
screen "02 Wip Select" 480x800, template "Current Menu Selection"
   Button "Top" at 375,164 size 100x101; TextOff 'Text'; PictureOff "basic panel top"
      on Press: function_b14e0dd5("pbs", 0)
      Appearance <- "[0]"
      Visibility <- "[0]"
   Button "Page Up" at 375,270 size 100x101; TextOff 'Text'; PictureOff "basic panel page up"
      on Press: function_b14e0dd5("pbs", 1)
      Visibility <- "[1]"
      Appearance <- "[1]"
   Button "Line Up" at 375,376 size 100x101; TextOff 'Text'; PictureOff "basic panel line up"
      on Press: function_b14e0dd5("pbs", 2)
      Appearance <- "[2]"
      Visibility <- "[2]"
   Button "Line Down" at 375,482 size 100x101; TextOff 'Text'; PictureOff "basic panel line down"
      on Press: function_b14e0dd5("pbs", 3)
      Visibility <- "[3]"
      Appearance <- "[3]"
   Button "Page Down" at 375,588 size 100x101; TextOff 'Text'; PictureOff "basic panel page down"
      on Press: function_b14e0dd5("pbs", 4)
      Appearance <- "[4]"
      Visibility <- "[4]"
   Button "Bottom" at 375,694 size 100x101; TextOff 'Text'; PictureOff "basic panel bottom"
      on Press: function_b14e0dd5("pbs", 5)
      Visibility <- "[5]"
      Appearance <- "[5]"
   IOField "brdrShortR00" at 5,164 size 365x101; FormatPattern 1
      Visibility <- "[6]"
      Appearance <- "[6]"
   IOField "brdrShortR01" at 5,270 size 365x101; FormatPattern 1
      Visibility <- "[7]"
      Appearance <- "[7]"
   IOField "brdrShortR02" at 5,376 size 365x101; FormatPattern 1
      Visibility <- "[8]"
      Appearance <- "[8]"
   IOField "brdrShortR03" at 5,482 size 365x101; FormatPattern 1
      Visibility <- "[9]"
      Appearance <- "[9]"
   IOField "brdrShortR04" at 5,588 size 365x101; FormatPattern 1
      Visibility <- "[10]"
      Appearance <- "[10]"
   IOField "brdrShortR05" at 5,694 size 365x101; FormatPattern 1
      Visibility <- "[11]"
      Appearance <- "[11]"
   Button "pbShortSelectR00" at 5,164 size 365x101; TextOff 'Text'
      on Release: ActivateScreen("01 Part Select", 0)
      on Press: function_b14e0dd5("pbs", 6)
   Button "pbShortSelectR01" at 5,270 size 365x101; TextOff 'Text'
      on Release: ActivateScreen("01 Part Select", 0)
      on Press: function_b14e0dd5("pbs", 7)
   Button "pbShortSelectR02" at 5,376 size 365x101; TextOff 'Text'
      on Release: ActivateScreen("01 Part Select", 0)
      on Press: function_b14e0dd5("pbs", 8)
   Button "pbShortSelectR03" at 5,482 size 365x101; TextOff 'Text'
      on Release: ActivateScreen("01 Part Select", 0)
      on Press: function_b14e0dd5("pbs", 9)
   Button "pbShortSelectR04" at 5,588 size 365x101; TextOff 'Text'
      on Release: ActivateScreen("01 Part Select", 0)
      on Press: function_b14e0dd5("pbs", 10)
   Button "pbShortSelectR05" at 5,694 size 365x101; TextOff 'Text'
      on Release: ActivateScreen("01 Part Select", 0)
      on Press: function_b14e0dd5("pbs", 11)
   IOField "brdrLongR00" at 5,164 size 470x101; FormatPattern 1
      Visibility <- "[18]"
   IOField "brdrLongR01" at 5,270 size 470x101; FormatPattern 1
      Visibility <- "[19]"
   IOField "brdrLongR02" at 5,376 size 470x101; FormatPattern 1
      Visibility <- "[20]"
   IOField "brdrLongR03" at 5,482 size 470x101; FormatPattern 1
      Visibility <- "[21]"
   IOField "brdrLongR04" at 5,588 size 470x101; FormatPattern 1
      Visibility <- "[22]"
   IOField "brdrLongR05" at 5,694 size 470x101; FormatPattern 1
      Visibility <- "[23]"
   Button "pbLongtSelectR00" at 5,164 size 470x101; TextOff 'Text'
      on Release: ActivateScreen("01 Part Select", 0)
      on Press: function_b14e0dd5("pbs", 6)
      Visibility <- "[18]"
   Button "pbLongtSelectR01" at 5,270 size 470x101; TextOff 'Text'
      on Release: ActivateScreen("01 Part Select", 0)
      on Press: function_b14e0dd5("pbs", 7)
      Visibility <- "[19]"
   Button "pbLongtSelectR02" at 5,376 size 470x101; TextOff 'Text'
      on Release: ActivateScreen("01 Part Select", 0)
      on Press: function_b14e0dd5("pbs", 8)
      Visibility <- "[20]"
   Button "pbLongtSelectR03" at 5,482 size 470x101; TextOff 'Text'
      on Release: ActivateScreen("01 Part Select", 0)
      on Press: function_b14e0dd5("pbs", 9)
      Visibility <- "[21]"
   Button "pbLongtSelectR04" at 5,588 size 470x101; TextOff 'Text'
      on Release: ActivateScreen("01 Part Select", 0)
      on Press: function_b14e0dd5("pbs", 10)
      Visibility <- "[22]"
   Button "pbLongtSelectR05" at 5,694 size 470x101; TextOff 'Text'
      on Release: ActivateScreen("01 Part Select", 0)
      on Press: function_b14e0dd5("pbs", 11)
      Visibility <- "[23]"
   IOField "iofLongtMenuSelectR00" at 42,166 size 430x97; FormatPattern ????????????????????????????????????????????????????????????
      Visibility <- "[18]"
      Appearance <- "[18]"
      ProcessValue <- "[7]"
   IOField "iofLongtMenuSelectR01" at 42,272 size 430x97; FormatPattern ????????????????????????????????????????????????????????????
      Visibility <- "[19]"
      Appearance <- "[19]"
      ProcessValue <- "[9]"
   IOField "iofLongtMenuSelectR02" at 42,378 size 430x97; FormatPattern ????????????????????????????????????????????????????????????
      Visibility <- "[20]"
      Appearance <- "[20]"
      ProcessValue <- "[11]"
   IOField "iofLongtMenuSelectR03" at 42,484 size 430x97; FormatPattern ????????????????????????????????????????????????????????????
      Visibility <- "[21]"
      Appearance <- "[21]"
      ProcessValue <- "[13]"
   IOField "iofLongtMenuSelectR04" at 42,590 size 430x97; FormatPattern ????????????????????????????????????????????????????????????
      Visibility <- "[22]"
      Appearance <- "[22]"
      ProcessValue <- "[15]"
   IOField "iofLongtMenuSelectR05" at 42,696 size 430x97; FormatPattern ????????????????????????????????????????????????????????????
      Visibility <- "[23]"
      Appearance <- "[23]"
      ProcessValue <- "[17]"
   IOField "iofLongLabelR00" at 7,166 size 35x97; FormatPattern ????????????????????????????????????????
      Visibility <- "[18]"
      Appearance <- "[18]"
      ProcessValue <- "[6]"
   IOField "iofLongLabelR01" at 7,272 size 35x97; FormatPattern ????????????????????????????????????????
      Appearance <- "[19]"
      Visibility <- "[19]"
      ProcessValue <- "[8]"
   IOField "iofLongLabelR02" at 7,378 size 35x97; FormatPattern ????????????????????????????????????????
      Appearance <- "[20]"
      Visibility <- "[20]"
      ProcessValue <- "[10]"
   IOField "iofLongLabelR03" at 7,484 size 35x97; FormatPattern ????????????????????????????????????????
      Appearance <- "[21]"
      Visibility <- "[21]"
      ProcessValue <- "[12]"
   IOField "iofLongLabelR04" at 7,590 size 35x97; FormatPattern ????????????????????????????????????????
      Visibility <- "[22]"
      Appearance <- "[22]"
      ProcessValue <- "[14]"
   IOField "iofLongtLabelR05" at 7,696 size 35x97; FormatPattern ????????????????????????????????????????
      Appearance <- "[23]"
      Visibility <- "[23]"
      ProcessValue <- "[16]"
   IOField "iofShortMenuSelectR00" at 42,166 size 325x97; FormatPattern ????????????????????????????????????????????????????????????
      Visibility <- "[6]"
      Appearance <- "[6]"
      ProcessValue <- "[7]"
   IOField "iofShortMenuSelectR01" at 42,272 size 325x97; FormatPattern ????????????????????????????????????????????????????????????
      Visibility <- "[7]"
      Appearance <- "[7]"
      ProcessValue <- "[9]"
   IOField "iofShortMenuSelectR02" at 42,378 size 325x97; FormatPattern ????????????????????????????????????????????????????????????
      Visibility <- "[8]"
      Appearance <- "[8]"
      ProcessValue <- "[11]"
   IOField "iofShortMenuSelectR03" at 42,484 size 325x97; FormatPattern ????????????????????????????????????????????????????????????
      Visibility <- "[9]"
      Appearance <- "[9]"
      ProcessValue <- "[13]"
   IOField "iofShortMenuSelectR04" at 42,590 size 325x97; FormatPattern ????????????????????????????????????????????????????????????
      Visibility <- "[10]"
      Appearance <- "[10]"
      ProcessValue <- "[15]"
   IOField "iofShortMenuSelectR05" at 42,696 size 325x97; FormatPattern ????????????????????????????????????????????????????????????
      Visibility <- "[11]"
      Appearance <- "[11]"
      ProcessValue <- "[17]"
   IOField "iofShortLabelR00" at 7,166 size 35x97; FormatPattern ????????????????????????????????????????
      Appearance <- "[6]"
      Visibility <- "[6]"
      ProcessValue <- "[6]"
   IOField "iofShortLabelR01" at 7,272 size 35x97; FormatPattern ????????????????????????????????????????
      Appearance <- "[7]"
      Visibility <- "[7]"
      ProcessValue <- "[8]"
   IOField "iofShortLabelR02" at 7,378 size 35x97; FormatPattern ????????????????????????????????????????
      Appearance <- "[8]"
      Visibility <- "[8]"
      ProcessValue <- "[10]"
   IOField "iofShortLabelR03" at 7,484 size 35x97; FormatPattern ????????????????????????????????????????
      Appearance <- "[9]"
      Visibility <- "[9]"
      ProcessValue <- "[12]"
   IOField "iofShortLabelR04" at 7,590 size 35x97; FormatPattern ????????????????????????????????????????
      Appearance <- "[10]"
      Visibility <- "[10]"
      ProcessValue <- "[14]"
   IOField "iofShorttLabelR05" at 7,696 size 35x97; FormatPattern ????????????????????????????????????????
      Appearance <- "[11]"
      Visibility <- "[11]"
      ProcessValue <- "[16]"

Template "Current Menu Selection" 480x800
   IOField "Menu Select Label" at 6,5 size 470x154; FormatPattern ????????????????????????????????????????????????????????????
      Appearance <- "[0]"
      Visibility <- "[0]"
      ProcessValue <- "[0]"
   Button "PB Menu Select" at 6,5 size 470x154; TextOff 'Text'
      on Release: ActivateScreen("02 Wip Select", 0)
      on Press: function_b14e0dd5("pb", 0)
*)

(* ===== HMI "HMI_RT_7" =====
system functions are stored by id; their names below are inferred from use
connection "pc01": ETHERNET, SMART_S7_1500_OMS

HMI tags "Default tag table"
   "station" : HMI Station: Compressed = PLC "HMI Stations: HMI Data".me[4] AT %DB1.DBW0, 100 ms

screen "01 Part Select" 480x800, template "Current Menu Selection"
   Button "B7" at 6,164 size 233x154; TextOff 'Text'
      on Press: function_b14e0dd5("pbs", 7)
      Visibility <- "[7]"
   Button "B6" at 6,323 size 233x154; TextOff 'Text'
      on Press: function_b14e0dd5("pbs", 6)
      Visibility <- "[6]"
   Button "B5" at 6,482 size 233x154; TextOff 'Text'
      on Press: function_b14e0dd5("pbs", 5)
      Visibility <- "[5]"
   Button "B4" at 6,641 size 233x154; TextOff 'Text'
      on Press: function_b14e0dd5("pbs", 4)
      Visibility <- "[4]"
   Button "B3" at 244,164 size 232x154; TextOff 'Text'
      on Press: function_b14e0dd5("pbs", 3)
      Visibility <- "[3]"
   Button "B2" at 244,323 size 232x154; TextOff 'Text'
      on Press: function_b14e0dd5("pbs", 2)
      Visibility <- "[2]"
   Button "B1" at 244,482 size 232x154; TextOff 'Text'
      on Press: function_b14e0dd5("pbs", 1)
      Visibility <- "[1]"
   Button "B0" at 244,641 size 232x154; TextOff 'Text'
      on Press: function_b14e0dd5("pbs", 0)
   IOField "B7 Label" at 6,164 size 233x154; FormatPattern ????????????????????????????????????????
      Appearance <- "[7]"
      ProcessValue <- "[7]"
      Visibility <- "[7]"
   IOField "B6 Label" at 6,323 size 233x154; FormatPattern ????????????????????????????????????????
      Appearance <- "[6]"
      ProcessValue <- "[6]"
      Visibility <- "[6]"
   IOField "B5 Label" at 6,482 size 233x154; FormatPattern ????????????????????????????????????????
      Appearance <- "[5]"
      ProcessValue <- "[5]"
      Visibility <- "[5]"
   IOField "B4 Label" at 6,641 size 233x154; FormatPattern ????????????????????????????????????????
      Appearance <- "[4]"
      ProcessValue <- "[4]"
      Visibility <- "[4]"
   IOField "B3 Label" at 244,164 size 232x154; FormatPattern ????????????????????????????????????????
      Appearance <- "[3]"
      ProcessValue <- "[3]"
      Visibility <- "[3]"
   IOField "B2 Label" at 244,323 size 232x154; FormatPattern ????????????????????????????????????????
      Appearance <- "[2]"
      ProcessValue <- "[2]"
      Visibility <- "[2]"
   IOField "B1 Label" at 244,482 size 232x154; FormatPattern ????????????????????????????????????????
      Appearance <- "[1]"
      ProcessValue <- "[1]"
      Visibility <- "[1]"
   IOField "B0 Label" at 244,641 size 232x154; FormatPattern ????????????????????????????????????????
      Appearance <- "[0]"
      ProcessValue <- "[0]"
      Visibility <- "[0]"

screen "02 Menu Select" 480x800, template "Current Menu Selection"
   Button "Top" at 375,164 size 100x101; TextOff 'Text'; PictureOff "basic panel top"
      on Press: function_b14e0dd5("pbs", 0)
      Appearance <- "[0]"
      Visibility <- "[0]"
   Button "Page Up" at 375,270 size 100x101; TextOff 'Text'; PictureOff "basic panel page up"
      on Press: function_b14e0dd5("pbs", 1)
      Visibility <- "[1]"
      Appearance <- "[1]"
   Button "Line Up" at 375,376 size 100x101; TextOff 'Text'; PictureOff "basic panel line up"
      on Press: function_b14e0dd5("pbs", 2)
      Appearance <- "[2]"
      Visibility <- "[2]"
   Button "Line Down" at 375,482 size 100x101; TextOff 'Text'; PictureOff "basic panel line down"
      on Press: function_b14e0dd5("pbs", 3)
      Visibility <- "[3]"
      Appearance <- "[3]"
   Button "Page Down" at 375,588 size 100x101; TextOff 'Text'; PictureOff "basic panel page down"
      on Press: function_b14e0dd5("pbs", 4)
      Appearance <- "[4]"
      Visibility <- "[4]"
   Button "Bottom" at 375,694 size 100x101; TextOff 'Text'; PictureOff "basic panel bottom"
      on Press: function_b14e0dd5("pbs", 5)
      Visibility <- "[5]"
      Appearance <- "[5]"
   IOField "brdrShortR00" at 5,164 size 365x101; FormatPattern 1
      Visibility <- "[6]"
      Appearance <- "[6]"
   IOField "brdrShortR01" at 5,270 size 365x101; FormatPattern 1
      Visibility <- "[7]"
      Appearance <- "[7]"
   IOField "brdrShortR02" at 5,376 size 365x101; FormatPattern 1
      Visibility <- "[8]"
      Appearance <- "[8]"
   IOField "brdrShortR03" at 5,482 size 365x101; FormatPattern 1
      Visibility <- "[9]"
      Appearance <- "[9]"
   IOField "brdrShortR04" at 5,588 size 365x101; FormatPattern 1
      Visibility <- "[10]"
      Appearance <- "[10]"
   IOField "brdrShortR05" at 5,694 size 365x101; FormatPattern 1
      Visibility <- "[11]"
      Appearance <- "[11]"
   Button "pbShortSelectR00" at 5,164 size 365x101; TextOff 'Text'
      on Release: ActivateScreen("01 Part Select", 0)
      on Press: function_b14e0dd5("pbs", 6)
   Button "pbShortSelectR01" at 5,270 size 365x101; TextOff 'Text'
      on Release: ActivateScreen("01 Part Select", 0)
      on Press: function_b14e0dd5("pbs", 7)
   Button "pbShortSelectR02" at 5,376 size 365x101; TextOff 'Text'
      on Release: ActivateScreen("01 Part Select", 0)
      on Press: function_b14e0dd5("pbs", 8)
   Button "pbShortSelectR03" at 5,482 size 365x101; TextOff 'Text'
      on Release: ActivateScreen("01 Part Select", 0)
      on Press: function_b14e0dd5("pbs", 9)
   Button "pbShortSelectR04" at 5,588 size 365x101; TextOff 'Text'
      on Release: ActivateScreen("01 Part Select", 0)
      on Press: function_b14e0dd5("pbs", 10)
   Button "pbShortSelectR05" at 5,694 size 365x101; TextOff 'Text'
      on Release: ActivateScreen("01 Part Select", 0)
      on Press: function_b14e0dd5("pbs", 11)
   IOField "brdrLongR00" at 5,164 size 470x101; FormatPattern 1
      Visibility <- "[18]"
   IOField "brdrLongR01" at 5,270 size 470x101; FormatPattern 1
      Visibility <- "[19]"
   IOField "brdrLongR02" at 5,376 size 470x101; FormatPattern 1
      Visibility <- "[20]"
   IOField "brdrLongR03" at 5,482 size 470x101; FormatPattern 1
      Visibility <- "[21]"
   IOField "brdrLongR04" at 5,588 size 470x101; FormatPattern 1
      Visibility <- "[22]"
   IOField "brdrLongR05" at 5,694 size 470x101; FormatPattern 1
      Visibility <- "[23]"
   Button "pbLongtSelectR00" at 5,164 size 470x101; TextOff 'Text'
      on Release: ActivateScreen("01 Part Select", 0)
      on Press: function_b14e0dd5("pbs", 6)
      Visibility <- "[18]"
   Button "pbLongtSelectR01" at 5,270 size 470x101; TextOff 'Text'
      on Release: ActivateScreen("01 Part Select", 0)
      on Press: function_b14e0dd5("pbs", 7)
      Visibility <- "[19]"
   Button "pbLongtSelectR02" at 5,376 size 470x101; TextOff 'Text'
      on Release: ActivateScreen("01 Part Select", 0)
      on Press: function_b14e0dd5("pbs", 8)
      Visibility <- "[20]"
   Button "pbLongtSelectR03" at 5,482 size 470x101; TextOff 'Text'
      on Release: ActivateScreen("01 Part Select", 0)
      on Press: function_b14e0dd5("pbs", 9)
      Visibility <- "[21]"
   Button "pbLongtSelectR04" at 5,588 size 470x101; TextOff 'Text'
      on Release: ActivateScreen("01 Part Select", 0)
      on Press: function_b14e0dd5("pbs", 10)
      Visibility <- "[22]"
   Button "pbLongtSelectR05" at 5,694 size 470x101; TextOff 'Text'
      on Release: ActivateScreen("01 Part Select", 0)
      on Press: function_b14e0dd5("pbs", 11)
      Visibility <- "[23]"
   IOField "iofLongtMenuSelectR00" at 42,166 size 430x97; FormatPattern ????????????????????????????????????????????????????????????
      Visibility <- "[18]"
      ProcessValue <- "[7]"
      Appearance <- "[18]"
   IOField "iofLongtMenuSelectR01" at 42,272 size 430x97; FormatPattern ????????????????????????????????????????????????????????????
      Visibility <- "[19]"
      ProcessValue <- "[9]"
      Appearance <- "[19]"
   IOField "iofLongtMenuSelectR02" at 42,378 size 430x97; FormatPattern ????????????????????????????????????????????????????????????
      Visibility <- "[20]"
      ProcessValue <- "[11]"
      Appearance <- "[20]"
   IOField "iofLongtMenuSelectR03" at 42,484 size 430x97; FormatPattern ????????????????????????????????????????????????????????????
      Visibility <- "[21]"
      ProcessValue <- "[13]"
      Appearance <- "[21]"
   IOField "iofLongtMenuSelectR04" at 42,590 size 430x97; FormatPattern ????????????????????????????????????????????????????????????
      Visibility <- "[22]"
      ProcessValue <- "[15]"
      Appearance <- "[22]"
   IOField "iofLongtMenuSelectR05" at 42,696 size 430x97; FormatPattern ????????????????????????????????????????????????????????????
      Visibility <- "[23]"
      ProcessValue <- "[17]"
      Appearance <- "[22]"
   IOField "iofLongLabelR00" at 7,166 size 35x97; FormatPattern ????????????????????????????????????????
      Visibility <- "[18]"
      ProcessValue <- "[6]"
      Appearance <- "[18]"
   IOField "iofLongLabelR01" at 7,272 size 35x97; FormatPattern ????????????????????????????????????????
      Appearance <- "[19]"
      ProcessValue <- "[8]"
      Visibility <- "[19]"
   IOField "iofLongLabelR02" at 7,378 size 35x97; FormatPattern ????????????????????????????????????????
      Appearance <- "[20]"
      ProcessValue <- "[10]"
      Visibility <- "[20]"
   IOField "iofLongLabelR03" at 7,484 size 35x97; FormatPattern ????????????????????????????????????????
      Appearance <- "[21]"
      ProcessValue <- "[12]"
      Visibility <- "[21]"
   IOField "iofLongLabelR04" at 7,590 size 35x97; FormatPattern ????????????????????????????????????????
      Visibility <- "[22]"
      ProcessValue <- "[14]"
      Appearance <- "[22]"
   IOField "iofLongtLabelR05" at 7,696 size 35x97; FormatPattern ????????????????????????????????????????
      Appearance <- "[23]"
      ProcessValue <- "[16]"
      Visibility <- "[23]"
   IOField "iofShortMenuSelectR00" at 42,166 size 325x97; FormatPattern ????????????????????????????????????????????????????????????
      Visibility <- "[6]"
      ProcessValue <- "[7]"
      Appearance <- "[6]"
   IOField "iofShortMenuSelectR01" at 42,272 size 325x97; FormatPattern ????????????????????????????????????????????????????????????
      Visibility <- "[7]"
      ProcessValue <- "[9]"
      Appearance <- "[7]"
   IOField "iofShortMenuSelectR02" at 42,378 size 325x97; FormatPattern ????????????????????????????????????????????????????????????
      Visibility <- "[8]"
      ProcessValue <- "[11]"
      Appearance <- "[8]"
   IOField "iofShortMenuSelectR03" at 42,484 size 325x97; FormatPattern ????????????????????????????????????????????????????????????
      Visibility <- "[9]"
      ProcessValue <- "[13]"
      Appearance <- "[9]"
   IOField "iofShortMenuSelectR04" at 42,590 size 325x97; FormatPattern ????????????????????????????????????????????????????????????
      Visibility <- "[10]"
      ProcessValue <- "[15]"
      Appearance <- "[10]"
   IOField "iofShortMenuSelectR05" at 42,696 size 325x97; FormatPattern ????????????????????????????????????????????????????????????
      Visibility <- "[11]"
      ProcessValue <- "[17]"
      Appearance <- "[11]"
   IOField "iofShortLabelR00" at 7,166 size 35x97; FormatPattern ????????????????????????????????????????
      Appearance <- "[6]"
      ProcessValue <- "[6]"
      Visibility <- "[6]"
   IOField "iofShortLabelR01" at 7,272 size 35x97; FormatPattern ????????????????????????????????????????
      Appearance <- "[7]"
      ProcessValue <- "[8]"
      Visibility <- "[7]"
   IOField "iofShortLabelR02" at 7,378 size 35x97; FormatPattern ????????????????????????????????????????
      Appearance <- "[8]"
      ProcessValue <- "[10]"
      Visibility <- "[8]"
   IOField "iofShortLabelR03" at 7,484 size 35x97; FormatPattern ????????????????????????????????????????
      Appearance <- "[9]"
      ProcessValue <- "[12]"
      Visibility <- "[9]"
   IOField "iofShortLabelR04" at 7,590 size 35x97; FormatPattern ????????????????????????????????????????
      Appearance <- "[10]"
      ProcessValue <- "[14]"
      Visibility <- "[10]"
   IOField "iofShorttLabelR05" at 7,696 size 35x97; FormatPattern ????????????????????????????????????????
      Appearance <- "[11]"
      ProcessValue <- "[16]"
      Visibility <- "[11]"

Template "Current Menu Selection" 480x800
   IOField "Menu Select Label" at 6,5 size 470x154; FormatPattern ????????????????????????????????????????????????????????????
      Appearance <- "[0]"
      Visibility <- "[0]"
      ProcessValue <- "[0]"
   Button "PB Menu Select" at 6,5 size 470x154; TextOff 'Text'
      on Release: ActivateScreen("02 Menu Select", 0)
      on Press: function_b14e0dd5("pb", 0)
*)

(* ===== HMI "HMI_RT_1" =====
system functions are stored by id; their names below are inferred from use

ScreenModuleEditorView "Table Row" 1312x52
   TextField "tfLine" at 5,1 size 216x48; Text 'Text'
      Visibility <- "interface.tfLine.animate"
      Appearance <- "interface.tfLine.animate"
   TextField "tfTime" at 1085,1 size 222x48; Text 'Text'
      Visibility <- "interface.tfTime.animate"
      Appearance <- "interface.tfTime.animate"
   TextField "tfDropZone" at 211,1 size 236x48; Text 'Text'
      Visibility <- "interface.tfDropZone.animate"
      Appearance <- "interface.tfDropZone.animate"
   TextField "tfSLPartNumber" at 445,1 size 650x48; Text 'Text'
      Visibility <- "interface.tfPartNumber.animateSL"
      Appearance <- "interface.tfPartNumber.animateSL"
   Button "pbSelect" at 0,0 size 1312x52; TextOff 'Text'
      on Release: ResetBit("interface.pbSelection.actuate")
      on Press: SetBit("interface.pbSelection.actuate")
      Appearance <- "interface.pbSelection.animate"
      Visibility <- "interface.pbSelection.animate"
      ObjectEnable <- "interface.pbSelection.animate"
   Rectangle "rtBackground" at 0,0 size 1312x52
      Visibility <- "interface.rtBackground.animate"
      Appearance <- "interface.rtBackground.animate"
   TextField "tfDLPartNumber" at 445,1 size 650x48; Text 'Text'
      Visibility <- "interface.tfPartNumber.animateDL"
      Appearance <- "interface.tfPartNumber.animateDL"
*)

(* ===== HMI "HMI_RT_1" =====
system functions are stored by id; their names below are inferred from use

ScreenModuleEditorView "IO Field: Double Width: Stacked" 370x111
   IOField "tfLable" at 0,55 size 370x56; FormatPattern ????????????????????????????????????????
      on OnFinishInput: SetBit("Interface.inputFinished")
      Appearance <- "Interface.animate"
      Visibility <- "Interface.animate"
      ProcessValue <- "Interface.value"
      ObjectEnable <- "Interface.animate"
   TextField "iofData" at 0,0 size 370x55; Text 'Text'
*)

(* ===== HMI "HMI_RT_1" =====
system functions are stored by id; their names below are inferred from use

ScreenModuleEditorView "IO Field: Single Width; Stacked" 370x111
   IOField "tfLable" at 0,55 size 370x56; FormatPattern ????????????????????????????????????????
      on OnFinishInput: SetBit("Interface.inputFinished")
      Appearance <- "Interface.animate"
      Visibility <- "Interface.animate"
      ObjectEnable <- "Interface.animate"
      ProcessValue <- "Interface.value"
   TextField "iofData" at 0,0 size 370x55; Text 'Text'
*)

(* ===== HMI "HMI_RT_1" =====
system functions are stored by id; their names below are inferred from use

ScreenModuleEditorView "IO Field: Single Width; Stacked" 178x111
   IOField "tfLable" at 0,55 size 178x56; FormatPattern ????????????????????????????????????????
      on OnFinishInput: SetBit("Interface.inputFinished")
      Appearance <- "Interface.animate"
      Visibility <- "Interface.animate"
      ProcessValue <- "Interface.value"
      ObjectEnable <- "Interface.animate"
   TextField "iofData" at 0,0 size 178x55; Text 'Text'
*)

(* ===== HMI "HMI_RT_1" =====

ScreenModuleEditorView "Settings Station Row" 671x200
   TextField "tfLine" at 0,0 size 135x200; Text 'VOLVO 00'
   TextField "tfDropzone" at 135,0 size 40x200; Text '00'
   TextField "tfWIP" at 175,0 size 40x200; Text '00'
   Group "rowBtn00" at 215,0 size 456x25
   Group "rowBtn01" at 215,25 size 456x25
   Group "rowBtn02" at 215,50 size 456x25
   Group "rowBtn03" at 215,75 size 456x25
   Group "rowBtn04" at 215,100 size 456x25
   Group "rowBtn05" at 215,125 size 456x25
   Group "rowBtn06" at 215,150 size 456x25
   Group "rowBtn07" at 215,175 size 456x25
   TextField "tfLablBtn00" at 215,0 size 40x25; Text '00'
   TextField "tfAllottedBtn00" at 255,0 size 80x25; Text '00:00'
   TextField "tfCriticalBtn00" at 335,0 size 80x25; Text '00:00'
   TextField "tfPartNumberBtn00" at 415,0 size 256x25; Text '00.00.000.000.0000'
   TextField "tfLablBtn01" at 215,25 size 40x25; Text '00'
   TextField "tfAllottedBtn01" at 255,25 size 80x25; Text '00:00'
   TextField "tfCriticalBtn01" at 335,25 size 80x25; Text '00:00'
   TextField "tfPartNumberBtn01" at 415,25 size 256x25; Text '00.00.000.000.0000'
   TextField "tfLablBtn02" at 215,50 size 40x25; Text '00'
   TextField "tfAllottedBtn02" at 255,50 size 80x25; Text '00:00'
   TextField "tfCriticalBtn02" at 335,50 size 80x25; Text '00:00'
   TextField "tfPartNumberBtn02" at 415,50 size 256x25; Text '00.00.000.000.0000'
   TextField "tfLablBtn03" at 215,75 size 40x25; Text '00'
   TextField "tfAllottedBtn03" at 255,75 size 80x25; Text '00:00'
   TextField "tfCriticalBtn03" at 335,75 size 80x25; Text '00:00'
   TextField "tfPartNumberBtn03" at 415,75 size 256x25; Text '00.00.000.000.0000'
   TextField "tfLablBtn04" at 215,100 size 40x25; Text '00'
   TextField "tfAllottedBtn04" at 255,100 size 80x25; Text '00:00'
   TextField "tfCriticalBtn04" at 335,100 size 80x25; Text '00:00'
   TextField "tfPartNumberBtn04" at 415,100 size 256x25; Text '00.00.000.000.0000'
   TextField "tfLablBtn05" at 215,125 size 40x25; Text '00'
   TextField "tfAllottedBtn05" at 255,125 size 80x25; Text '00:00'
   TextField "tfCriticalBtn05" at 335,125 size 80x25; Text '00:00'
   TextField "tfPartNumberBtn05" at 415,125 size 256x25; Text '00.00.000.000.0000'
   TextField "tfLablBtn06" at 215,150 size 40x25; Text '00'
   TextField "tfAllottedBtn06" at 255,150 size 80x25; Text '00:00'
   TextField "tfCriticalBtn06" at 335,150 size 80x25; Text '00:00'
   TextField "tfPartNumberBtn06" at 415,150 size 256x25; Text '00.00.000.000.0000'
   TextField "tfLablBtn07" at 215,175 size 40x25; Text '00'
   TextField "tfAllottedBtn07" at 255,175 size 80x25; Text '00:00'
   TextField "tfCriticalBtn07" at 335,175 size 80x25; Text '00:00'
   TextField "tfPartNumberBtn07" at 415,175 size 256x25; Text '00.00.000.000.0000'
*)

(* ===== HMI "HMI_RT_1" =====

ScreenModuleEditorView "Settings Station Row" 671x200
   TextField "tfLine" at 0,0 size 135x200; Text 'VOLVO 00'
   TextField "tfDropzone" at 135,0 size 40x200; Text '00'
   TextField "tfWIP" at 175,0 size 40x200; Text '00'
   Group "rowBtn00" at 215,0 size 456x25
   Group "rowBtn01" at 215,25 size 456x25
   Group "rowBtn02" at 215,50 size 456x25
   Group "rowBtn03" at 215,75 size 456x25
   Group "rowBtn04" at 215,100 size 456x25
   Group "rowBtn05" at 215,125 size 456x25
   Group "rowBtn06" at 215,150 size 456x25
   Group "rowBtn07" at 215,175 size 456x25
   TextField "tfLablBtn00" at 215,0 size 40x25; Text '00'
   TextField "tfAllottedBtn00" at 255,0 size 80x25; Text '00:00'
   TextField "tfCriticalBtn00" at 335,0 size 80x25; Text '00:00'
   TextField "tfPartNumberBtn00" at 415,0 size 256x25; Text '00.00.000.000.0000'
   TextField "tfLablBtn01" at 215,25 size 40x25; Text '00'
   TextField "tfAllottedBtn01" at 255,25 size 80x25; Text '00:00'
   TextField "tfCriticalBtn01" at 335,25 size 80x25; Text '00:00'
   TextField "tfPartNumberBtn01" at 415,25 size 256x25; Text '00.00.000.000.0000'
   TextField "tfLablBtn02" at 215,50 size 40x25; Text '00'
   TextField "tfAllottedBtn02" at 255,50 size 80x25; Text '00:00'
   TextField "tfCriticalBtn02" at 335,50 size 80x25; Text '00:00'
   TextField "tfPartNumberBtn02" at 415,50 size 256x25; Text '00.00.000.000.0000'
   TextField "tfLablBtn03" at 215,75 size 40x25; Text '00'
   TextField "tfAllottedBtn03" at 255,75 size 80x25; Text '00:00'
   TextField "tfCriticalBtn03" at 335,75 size 80x25; Text '00:00'
   TextField "tfPartNumberBtn03" at 415,75 size 256x25; Text '00.00.000.000.0000'
   TextField "tfLablBtn04" at 215,100 size 40x25; Text '00'
   TextField "tfAllottedBtn04" at 255,100 size 80x25; Text '00:00'
   TextField "tfCriticalBtn04" at 335,100 size 80x25; Text '00:00'
   TextField "tfPartNumberBtn04" at 415,100 size 256x25; Text '00.00.000.000.0000'
   TextField "tfLablBtn05" at 215,125 size 40x25; Text '00'
   TextField "tfAllottedBtn05" at 255,125 size 80x25; Text '00:00'
   TextField "tfCriticalBtn05" at 335,125 size 80x25; Text '00:00'
   TextField "tfPartNumberBtn05" at 415,125 size 256x25; Text '00.00.000.000.0000'
   TextField "tfLablBtn06" at 215,150 size 40x25; Text '00'
   TextField "tfAllottedBtn06" at 255,150 size 80x25; Text '00:00'
   TextField "tfCriticalBtn06" at 335,150 size 80x25; Text '00:00'
   TextField "tfPartNumberBtn06" at 415,150 size 256x25; Text '00.00.000.000.0000'
   TextField "tfLablBtn07" at 215,175 size 40x25; Text '00'
   TextField "tfAllottedBtn07" at 255,175 size 80x25; Text '00:00'
   TextField "tfCriticalBtn07" at 335,175 size 80x25; Text '00:00'
   TextField "tfPartNumberBtn07" at 415,175 size 256x25; Text '00.00.000.000.0000'
*)

(* ===== HMI "HMI_RT_1" =====

ScreenModuleEditorView "Settings Station Row" 671x200
   TextField "tfLine" at 0,0 size 135x200; Text 'VOLVO 00'
   TextField "tfDropzone" at 135,0 size 40x200; Text '00'
   TextField "tfWIP" at 175,0 size 40x200; Text '00'
   Group "rowBtn00" at 215,0 size 456x25
   Group "rowBtn01" at 215,25 size 456x25
   Group "rowBtn02" at 215,50 size 456x25
   Group "rowBtn03" at 215,75 size 456x25
   Group "rowBtn04" at 215,100 size 456x25
   Group "rowBtn05" at 215,125 size 456x25
   Group "rowBtn06" at 215,150 size 456x25
   Group "rowBtn07" at 215,175 size 456x25
   TextField "tfLablBtn00" at 215,0 size 40x25; Text '00'
   TextField "tfAllottedBtn00" at 255,0 size 80x25; Text '00:00'
   TextField "tfCriticalBtn00" at 335,0 size 80x25; Text '00:00'
   TextField "tfPartNumberBtn00" at 415,0 size 256x25; Text '00.00.000.000.0000'
   TextField "tfLablBtn01" at 215,25 size 40x25; Text '00'
   TextField "tfAllottedBtn01" at 255,25 size 80x25; Text '00:00'
   TextField "tfCriticalBtn01" at 335,25 size 80x25; Text '00:00'
   TextField "tfPartNumberBtn01" at 415,25 size 256x25; Text '00.00.000.000.0000'
   TextField "tfLablBtn02" at 215,50 size 40x25; Text '00'
   TextField "tfAllottedBtn02" at 255,50 size 80x25; Text '00:00'
   TextField "tfCriticalBtn02" at 335,50 size 80x25; Text '00:00'
   TextField "tfPartNumberBtn02" at 415,50 size 256x25; Text '00.00.000.000.0000'
   TextField "tfLablBtn03" at 215,75 size 40x25; Text '00'
   TextField "tfAllottedBtn03" at 255,75 size 80x25; Text '00:00'
   TextField "tfCriticalBtn03" at 335,75 size 80x25; Text '00:00'
   TextField "tfPartNumberBtn03" at 415,75 size 256x25; Text '00.00.000.000.0000'
   TextField "tfLablBtn04" at 215,100 size 40x25; Text '00'
   TextField "tfAllottedBtn04" at 255,100 size 80x25; Text '00:00'
   TextField "tfCriticalBtn04" at 335,100 size 80x25; Text '00:00'
   TextField "tfPartNumberBtn04" at 415,100 size 256x25; Text '00.00.000.000.0000'
   TextField "tfLablBtn05" at 215,125 size 40x25; Text '00'
   TextField "tfAllottedBtn05" at 255,125 size 80x25; Text '00:00'
   TextField "tfCriticalBtn05" at 335,125 size 80x25; Text '00:00'
   TextField "tfPartNumberBtn05" at 415,125 size 256x25; Text '00.00.000.000.0000'
   TextField "tfLablBtn06" at 215,150 size 40x25; Text '00'
   TextField "tfAllottedBtn06" at 255,150 size 80x25; Text '00:00'
   TextField "tfCriticalBtn06" at 335,150 size 80x25; Text '00:00'
   TextField "tfPartNumberBtn06" at 415,150 size 256x25; Text '00.00.000.000.0000'
   TextField "tfLablBtn07" at 215,175 size 40x25; Text '00'
   TextField "tfAllottedBtn07" at 255,175 size 80x25; Text '00:00'
   TextField "tfCriticalBtn07" at 335,175 size 80x25; Text '00:00'
   TextField "tfPartNumberBtn07" at 415,175 size 256x25; Text '00.00.000.000.0000'
*)

(* ===== HMI "HMI_RT_1" =====

ScreenModuleEditorView "Settings Station Row" 671x200
   TextField "tfLine" at 0,0 size 135x200; Text 'VOLVO 00'
   TextField "tfDropzone" at 135,0 size 40x200; Text '00'
   TextField "tfWIP" at 175,0 size 40x200; Text '00'
   TextField "tfLablBtn00" at 215,0 size 40x25; Text '00'
   TextField "tfAllottedBtn00" at 255,0 size 80x25; Text '00:00'
   TextField "tfCriticalBtn00" at 335,0 size 80x25; Text '00:00'
   TextField "tfPartNumberBtn00" at 415,0 size 256x25; Text '00.00.000.000.0000'
   TextField "tfLablBtn01" at 215,25 size 40x25; Text '00'
   TextField "tfAllottedBtn01" at 255,25 size 80x25; Text '00:00'
   TextField "tfCriticalBtn01" at 335,25 size 80x25; Text '00:00'
   TextField "tfPartNumberBtn01" at 415,25 size 256x25; Text '00.00.000.000.0000'
   TextField "tfLablBtn02" at 215,50 size 40x25; Text '00'
   TextField "tfAllottedBtn02" at 255,50 size 80x25; Text '00:00'
   TextField "tfCriticalBtn02" at 335,50 size 80x25; Text '00:00'
   TextField "tfPartNumberBtn02" at 415,50 size 256x25; Text '00.00.000.000.0000'
   TextField "tfLablBtn03" at 215,75 size 40x25; Text '00'
   TextField "tfAllottedBtn03" at 255,75 size 80x25; Text '00:00'
   TextField "tfCriticalBtn03" at 335,75 size 80x25; Text '00:00'
   TextField "tfPartNumberBtn03" at 415,75 size 256x25; Text '00.00.000.000.0000'
   TextField "tfLablBtn04" at 215,100 size 40x25; Text '00'
   TextField "tfAllottedBtn04" at 255,100 size 80x25; Text '00:00'
   TextField "tfCriticalBtn04" at 335,100 size 80x25; Text '00:00'
   TextField "tfPartNumberBtn04" at 415,100 size 256x25; Text '00.00.000.000.0000'
   TextField "tfLablBtn05" at 215,125 size 40x25; Text '00'
   TextField "tfAllottedBtn05" at 255,125 size 80x25; Text '00:00'
   TextField "tfCriticalBtn05" at 335,125 size 80x25; Text '00:00'
   TextField "tfPartNumberBtn05" at 415,125 size 256x25; Text '00.00.000.000.0000'
   TextField "tfLablBtn06" at 215,150 size 40x25; Text '00'
   TextField "tfAllottedBtn06" at 255,150 size 80x25; Text '00:00'
   TextField "tfCriticalBtn06" at 335,150 size 80x25; Text '00:00'
   TextField "tfPartNumberBtn06" at 415,150 size 256x25; Text '00.00.000.000.0000'
   TextField "tfLablBtn07" at 215,175 size 40x25; Text '00'
   TextField "tfAllottedBtn07" at 255,175 size 80x25; Text '00:00'
   TextField "tfCriticalBtn07" at 335,175 size 80x25; Text '00:00'
   TextField "tfPartNumberBtn07" at 415,175 size 256x25; Text '00.00.000.000.0000'
   TextField "tfPNDoubleBtn00" at 415,0 size 256x25; Text '00.00.000.000.0000 00.00.000.000.0000'
   TextField "tfPNDoubleBtn01" at 415,25 size 256x25; Text '00.00.000.000.0000 00.00.000.000.0000'
   TextField "tfPNDoubleBtn02" at 415,50 size 256x25; Text '00.00.000.000.0000 00.00.000.000.0000'
   TextField "tfPNDoubleBtn03" at 415,75 size 256x25; Text '00.00.000.000.0000 00.00.000.000.0000'
   TextField "tfPNDoubleBtn04" at 415,100 size 256x25; Text '00.00.000.000.0000 00.00.000.000.0000'
   TextField "tfPNDoubleBtn05" at 415,125 size 256x25; Text '00.00.000.000.0000 00.00.000.000.0000'
   TextField "tfPNDoubleBtn06" at 415,150 size 256x25; Text '00.00.000.000.0000 00.00.000.000.0000'
   TextField "tfPNDoubleBtn07" at 415,175 size 256x25; Text '00.00.000.000.0000 00.00.000.000.0000'
*)

(* ===== HMI "HMI_RT_1" =====

graphic list "Top": 0 '100 x 100 Top'; 1 '100 x 100 Actuated Top'

graphic list "Page Up": 0 '100 x 100 Page Up'; 1 '100 x 100 Actuated Page Up'

graphic list "Line Up": 0 '100 x 100 Line Up'; 1 '100 x 100 Actuated Line Up'

graphic list "Line Down": 0 '100 x 100 Line Down'; 1 '100 x 100 Actuated Line Down'

graphic list "Page Down": 0 '100 x 100 Page Down'; 1 '100 x 100 Actuated Page Down'

graphic list "Bottom": 0 '100 x 100 Bottom'; 1 '100 x 100 Actuated Bottom'

ScreenModuleEditorView "Nav Bar: Vertical" 100x600
   Button "btnTop" at 1,1 size 98x98; TextOff 'Text'; PictureList "Top"
   Button "btnPageUp" at 1,101 size 98x98; TextOff 'Text'; PictureList "Page Up"
   Button "btnLineUp" at 1,201 size 98x98; TextOff 'Text'; PictureList "Line Up"
   Button "btnLineDown" at 1,301 size 98x98; TextOff 'Text'; PictureList "Line Down"
   Button "btnPageDown" at 1,401 size 98x98; TextOff 'Text'; PictureList "Page Down"
   Button "btnBottom" at 1,501 size 98x98; TextOff 'Text'; PictureList "Bottom"
*)

(* ===== HMI "HMI_RT_1" =====
system functions are stored by id; their names below are inferred from use

graphic list "Top": 0 '100 x 100 Top'; 1 '100 x 100 Actuated Top'

graphic list "Page Up": 0 '100 x 100 Page Up'; 1 '100 x 100 Actuated Page Up'

graphic list "Line Up": 0 '100 x 100 Line Up'; 1 '100 x 100 Actuated Line Up'

graphic list "Line Down": 0 '100 x 100 Line Down'; 1 '100 x 100 Actuated Line Down'

graphic list "Page Down": 0 '100 x 100 Page Down'; 1 '100 x 100 Actuated Page Down'

graphic list "Bottom": 0 '100 x 100 Bottom'; 1 '100 x 100 Actuated Bottom'

ScreenModuleEditorView "Nav Bar: Vertical" 100x600
   Button "btnTop" at 1,1 size 98x98; TextOff 'Text'; PictureList "Top"
      on Press: SetBit("TableNavBar.top.actuate")
      on Release: ResetBit("TableNavBar.top.actuate")
      Visibility <- "TableNavBar.top.visible"
      ObjectEnable <- "TableNavBar.top.enable"
      ProcessValue <- "TableNavBar.top.listSelect"
      Appearance <- "TableNavBar.top.animate"
   Button "btnPageUp" at 1,101 size 98x98; TextOff 'Text'; PictureList "Page Up"
      on Release: ResetBit("TableNavBar.pageUp.actuate")
      on Press: SetBit("TableNavBar.pageUp.actuate")
      ProcessValue <- "TableNavBar.pageUp.listSelect"
      Appearance <- "TableNavBar.pageUp.animate"
      ObjectEnable <- "TableNavBar.pageUp.enable"
      Visibility <- "TableNavBar.pageUp.visible"
   Button "btnLineUp" at 1,201 size 98x98; TextOff 'Text'; PictureList "Line Up"
      on Release: ResetBit("TableNavBar.lineUp.actuate")
      on Press: SetBit("TableNavBar.lineUp.actuate")
      ProcessValue <- "TableNavBar.lineUp.listSelect"
      Visibility <- "TableNavBar.lineUp.visible"
      ObjectEnable <- "TableNavBar.lineUp.enable"
      Appearance <- "TableNavBar.lineUp.animate"
   Button "btnLineDown" at 1,301 size 98x98; TextOff 'Text'; PictureList "Line Down"
      on Release: ResetBit("TableNavBar.lineDown.actuate")
      on Press: SetBit("TableNavBar.lineDown.actuate")
      ProcessValue <- "TableNavBar.lineDown.listSelect"
      Appearance <- "TableNavBar.lineDown.animate"
      ObjectEnable <- "TableNavBar.lineDown.enable"
      Visibility <- "TableNavBar.lineDown.visible"
   Button "btnPageDown" at 1,401 size 98x98; TextOff 'Text'; PictureList "Page Down"
      on Release: ResetBit("TableNavBar.pageDown.actuate")
      on Press: SetBit("TableNavBar.pageDown.actuate")
      ProcessValue <- "TableNavBar.pageDown.listSelect"
      Visibility <- "TableNavBar.pageDown.visible"
      ObjectEnable <- "TableNavBar.pageDown.enable"
      Appearance <- "TableNavBar.pageDown.animate"
   Button "btnBottom" at 1,501 size 98x98; TextOff 'Text'; PictureList "Bottom"
      on Release: ResetBit("TableNavBar.bottom.actuate")
      on Press: SetBit("TableNavBar.bottom.actuate")
      ProcessValue <- "TableNavBar.bottom.listSelect"
      Appearance <- "TableNavBar.bottom.animate"
      ObjectEnable <- "TableNavBar.bottom.enable"
      Visibility <- "TableNavBar.bottom.visible"
*)

(* ===== HMI "HMI_RT_1" =====
system functions are stored by id; their names below are inferred from use

graphic list "Top": 0 '100 x 100 Top'; 1 '100 x 100 Actuated Top'

graphic list "Page Up": 0 '100 x 100 Page Up'; 1 '100 x 100 Actuated Page Up'

graphic list "Line Up": 0 '100 x 100 Line Up'; 1 '100 x 100 Actuated Line Up'

graphic list "Line Down": 0 '100 x 100 Line Down'; 1 '100 x 100 Actuated Line Down'

graphic list "Page Down": 0 '100 x 100 Page Down'; 1 '100 x 100 Actuated Page Down'

graphic list "Bottom": 0 '100 x 100 Bottom'; 1 '100 x 100 Actuated Bottom'

ScreenModuleEditorView "Nav Bar: Horizontal" 100x600
   Button "btnTop" at 1,1 size 98x98; TextOff 'Text'; PictureList "Top"
      on Release: ResetBit("TableNavBar.top.actuate")
      on Press: SetBit("TableNavBar.top.actuate")
      Visibility <- "TableNavBar.top.visible"
      ObjectEnable <- "TableNavBar.top.enable"
      ProcessValue <- "TableNavBar.top.listSelect"
      Appearance <- "TableNavBar.top.animate"
   Button "btnPageUp" at 1,101 size 98x98; TextOff 'Text'; PictureList "Page Up"
      on Release: ResetBit("TableNavBar.pageUp.actuate")
      on Press: SetBit("TableNavBar.pageUp.actuate")
      Appearance <- "TableNavBar.pageUp.animate"
      ObjectEnable <- "TableNavBar.pageUp.enable"
      ProcessValue <- "TableNavBar.pageUp.listSelect"
      Visibility <- "TableNavBar.pageUp.visible"
   Button "btnLineUp" at 1,201 size 98x98; TextOff 'Text'; PictureList "Line Up"
      on Release: ResetBit("TableNavBar.lineUp.actuate")
      on Press: SetBit("TableNavBar.lineUp.actuate")
      Visibility <- "TableNavBar.lineUp.visible"
      ObjectEnable <- "TableNavBar.lineUp.enable"
      ProcessValue <- "TableNavBar.lineUp.listSelect"
      Appearance <- "TableNavBar.lineUp.animate"
   Button "btnLineDown" at 1,301 size 98x98; TextOff 'Text'; PictureList "Line Down"
      on Release: ResetBit("TableNavBar.lineDown.actuate")
      on Press: SetBit("TableNavBar.lineDown.actuate")
      Appearance <- "TableNavBar.lineDown.animate"
      ObjectEnable <- "TableNavBar.lineDown.enable"
      ProcessValue <- "TableNavBar.lineDown.listSelect"
      Visibility <- "TableNavBar.lineDown.visible"
   Button "btnPageDown" at 1,401 size 98x98; TextOff 'Text'; PictureList "Page Down"
      on Release: ResetBit("TableNavBar.pageDown.actuate")
      on Press: SetBit("TableNavBar.pageDown.actuate")
      Visibility <- "TableNavBar.pageDown.visible"
      ObjectEnable <- "TableNavBar.pageDown.enable"
      ProcessValue <- "TableNavBar.pageDown.listSelect"
      Appearance <- "TableNavBar.pageDown.animate"
   Button "btnBottom" at 1,501 size 98x98; TextOff 'Text'; PictureList "Bottom"
      on Release: ResetBit("TableNavBar.bottom.actuate")
      on Press: SetBit("TableNavBar.bottom.actuate")
      Appearance <- "TableNavBar.bottom.animate"
      ObjectEnable <- "TableNavBar.bottom.enable"
      ProcessValue <- "TableNavBar.bottom.listSelect"
      Visibility <- "TableNavBar.bottom.visible"
*)

(* ===== HMI "HMI_RT_1" =====
system functions are stored by id; their names below are inferred from use

graphic list "Top": 0 '100 x 100 Top'; 1 '100 x 100 Actuated Top'

graphic list "Page Up": 0 '100 x 100 Page Up'; 1 '100 x 100 Actuated Page Up'

graphic list "Line Up": 0 '100 x 100 Line Up'; 1 '100 x 100 Actuated Line Up'

graphic list "Line Down": 0 '100 x 100 Line Down'; 1 '100 x 100 Actuated Line Down'

graphic list "Page Down": 0 '100 x 100 Page Down'; 1 '100 x 100 Actuated Page Down'

graphic list "Bottom": 0 '100 x 100 Bottom'; 1 '100 x 100 Actuated Bottom'

ScreenModuleEditorView "Nav Bar: Horizontal" 600x100
   Button "btnTop" at 1,1 size 98x98; TextOff 'Text'; PictureList "Top"
      on Release: ResetBit("TableNavBar.top.actuate")
      on Press: SetBit("TableNavBar.top.actuate")
      Visibility <- "TableNavBar.top.visible"
      ObjectEnable <- "TableNavBar.top.enable"
      ProcessValue <- "TableNavBar.top.listSelect"
      Appearance <- "TableNavBar.top.animate"
   Button "btnPageUp" at 101,1 size 98x98; TextOff 'Text'; PictureList "Page Up"
      on Release: ResetBit("TableNavBar.pageUp.actuate")
      on Press: SetBit("TableNavBar.pageUp.actuate")
      Appearance <- "TableNavBar.pageUp.animate"
      ObjectEnable <- "TableNavBar.pageUp.enable"
      ProcessValue <- "TableNavBar.pageUp.listSelect"
      Visibility <- "TableNavBar.pageUp.visible"
   Button "btnLineUp" at 201,1 size 98x98; TextOff 'Text'; PictureList "Line Up"
      on Release: ResetBit("TableNavBar.lineUp.actuate")
      on Press: SetBit("TableNavBar.lineUp.actuate")
      Visibility <- "TableNavBar.lineUp.visible"
      ObjectEnable <- "TableNavBar.lineUp.enable"
      ProcessValue <- "TableNavBar.lineUp.listSelect"
      Appearance <- "TableNavBar.lineUp.animate"
   Button "btnLineDown" at 301,1 size 98x98; TextOff 'Text'; PictureList "Line Down"
      on Release: ResetBit("TableNavBar.lineDown.actuate")
      on Press: SetBit("TableNavBar.lineDown.actuate")
      Appearance <- "TableNavBar.lineDown.animate"
      ObjectEnable <- "TableNavBar.lineDown.enable"
      ProcessValue <- "TableNavBar.lineDown.listSelect"
      Visibility <- "TableNavBar.lineDown.visible"
   Button "btnPageDown" at 401,1 size 98x98; TextOff 'Text'; PictureList "Page Down"
      on Release: ResetBit("TableNavBar.pageDown.actuate")
      on Press: SetBit("TableNavBar.pageDown.actuate")
      Visibility <- "TableNavBar.pageDown.visible"
      ObjectEnable <- "TableNavBar.pageDown.enable"
      ProcessValue <- "TableNavBar.pageDown.listSelect"
      Appearance <- "TableNavBar.pageDown.animate"
   Button "btnBottom" at 501,1 size 98x98; TextOff 'Text'; PictureList "Bottom"
      on Release: ResetBit("TableNavBar.bottom.actuate")
      on Press: SetBit("TableNavBar.bottom.actuate")
      Appearance <- "TableNavBar.bottom.animate"
      ObjectEnable <- "TableNavBar.bottom.enable"
      ProcessValue <- "TableNavBar.bottom.listSelect"
      Visibility <- "TableNavBar.bottom.visible"
*)

(* ===== HMI "HMI_RT_1" =====
system functions are stored by id; their names below are inferred from use

ScreenModuleEditorView "PB: Dynamic Text Label" 100x100
   Button "pbActuate" at 0,0 size 100x100; TextOff 'Text'
      on Press: SetBit("Interface.actuate")
      on Release: ResetBit("Interface.actuate")
      ObjectEnable <- "Interface.enable"
      Visibility <- "Interface.visible"
   TextField "tfDisplay" at 0,0 size 100x100; Text 'Text'
      Visibility <- "Interface.visible"
      Appearance <- "Interface.animate"
*)

(* ===== HMI "HMI_RT_1" =====
system functions are stored by id; their names below are inferred from use

ScreenModuleEditorView "PB: Static Text Label" 274x45
   Button "Select All Stations" at 0,0 size 274x45; TextOff 'Text'
      on Press: function_b14e0dd5("Interface.actuate", 0)
      Appearance <- "Interface.animate"
      ObjectEnable <- "Interface.animate"
      Visibility <- "Interface.animate"
*)

(* ===== HMI "HMI_RT_1" =====

